TYPE "HMI Station: Wip Select: Screen"
   STRUCT
      animate : Array[0.."wipSelScrnObjCnt"] of Int;
      pbs : DWord;
      txt : Array[0.."wipSelScrnObjCnt"] of WString ["LONG_STRING_LENGTH"];
   END_STRUCT;
   // // txt[6] : wip select 00 label
   // // txt[7] : wip select 00 text
   // // txt[8] : wip select 01 label
   // // txt[9] : wip select 01 text
   // // txt[10] : wip select 02 label
   // // txt[11] : wip select 02 text
   // // txt[12] : wip select 03 label
   // // txt[13] : wip select 03 text
   // // txt[14] : wip select 04 label
   // // txt[15] : wip select 04 text
   // // txt[16] : wip select 05 label
   // // txt[17] : wip select 05 text
END_TYPE

TYPE "HMI Station: Template Screen"
   STRUCT
      animate : Array[0.."tmpltScrnObjCnt"] of Int;
      pb : DWord;
      text : Array[0.."tmpltScrnObjCnt"] of WString ["LONG_STRING_LENGTH"];
   END_STRUCT;
END_TYPE

// folder: KP8 Driver

TYPE "KP8 I/O Data"
   STRUCT
      input : Word;
      tempOut : DWord;
      finalOut : DWord;
   END_STRUCT;
END_TYPE

TYPE "KP8 Driver: Parameters: 1 Button"
   STRUCT
      activate : Bool;   // true = button on, flase = button off
      cOn1 : String[10];   // color when button is in pressed state. valid entries: 'red', 'green', 'blue', 'yellow', 'white', 'off'
      cOn2 : String[10];   // second flash color when button is pressed and flashing is enabled. valid entries: 'red', 'green', 'blue', 'yellow', 'white', 'off'
      cOff : String[10];   // color when button is in un-pressed state. valid entries: 'red', 'green', 'blue', 'yellow', 'white', 'off'
      flash : Bool;   // false = color 1, true = color 2. set to clock bit to flash at that rate
      group : Int;   // 0 disables. buttons in groups have a mutually exclusive 'on' state.
      mode : Bool;   // true = maintained, fales = momentary
   END_STRUCT;
END_TYPE

TYPE "KP8 Driver: Button States"
   STRUCT
      btn : Array[0..7] of Bool;
   END_STRUCT;
END_TYPE

TYPE "KP8 Driver: Parameters: 8 Buttons"
   STRUCT
      btn : Array[0..7] of "KP8 Driver: Parameters: 1 Button";
   END_STRUCT;
END_TYPE

TYPE "KP8 Driver: Feedback Data"
   STRUCT
      acutal : "KP8 Driver: Button States";
      falling : "KP8 Driver: Button States";
      rising : "KP8 Driver: Button States";
   END_STRUCT;
END_TYPE

// folder: Linked List

TYPE "Linked List: Node: Data"
   STRUCT
      place_holder : Int;
   END_STRUCT;
END_TYPE

TYPE "Linked List: Node: Meta"
   STRUCT
      key : DInt := -1;
      is_head : Bool;
      is_tail : Bool;
      next : DInt := -1;
   END_STRUCT;
END_TYPE

TYPE "Linked List: Node"
   STRUCT
      data : "Linked List: Node: Data";
      meta : "Linked List: Node: Meta";
   END_STRUCT;
END_TYPE

TYPE "Linked List: List"
   STRUCT
      me : Array[0.."LINKED_LIST_LENGTH"] of "Linked List: Node";
   END_STRUCT;
END_TYPE

TYPE "Linked List: Method Interface: Reset: In"
   STRUCT
      request : Bool;
   END_STRUCT;
END_TYPE

TYPE "Linked List: Method Interface: Reverse: Out"
   STRUCT
      done : Bool;
      error : Bool;
      error_message : String;
   END_STRUCT;
END_TYPE

TYPE "Linked List: Method Interface: Reverse: In"
   STRUCT
      request : Bool;
   END_STRUCT;
END_TYPE

TYPE "Linked List: Method Interface: Display: Out"
   STRUCT
      done : Bool;
      list : "Linked List: List";
   END_STRUCT;
END_TYPE

TYPE "Linked List: Method Interface: Display: In"
   STRUCT
      request : Bool;
   END_STRUCT;
END_TYPE

TYPE "Linked List: Method Interface: Search: Out"
   STRUCT
      done : Bool;
      error : Bool;
      error_message : String;
      found : Bool;
      not_found : Bool;
      returned_node : "Linked List: Node";
   END_STRUCT;
END_TYPE

TYPE "Linked List: Method Interface: Search: In"
   STRUCT
      data : "Linked List: Node: Data";
      request : Bool;
   END_STRUCT;
END_TYPE

TYPE "Linked List: Method Interface: Reset: Out"
   STRUCT
      done : Bool;
   END_STRUCT;
END_TYPE

TYPE "Linked List: Method Interface: Delete: Out"
   STRUCT
      done : Bool;
      error : Bool;
      error_message : String;
   END_STRUCT;
END_TYPE

TYPE "Linked List: Method Interface: Delete: In"
   STRUCT
      node : "Linked List: Node";   // key of node to be deleted
      request : Bool;
   END_STRUCT;
END_TYPE

TYPE "Linked List: Method Interface: Insert: Out"
   STRUCT
      done : Bool;
      error : Bool;
      error_message : String;
   END_STRUCT;
END_TYPE

TYPE "Linked List: Method Interface: Insert: In"
   STRUCT
      target_node : "Linked List: Node";   // key of node after which new node is to be inserted
      data : "Linked List: Node: Data";
      request : Bool;
   END_STRUCT;
END_TYPE

TYPE "Linked List: Method Interface: Append: In"
   STRUCT
      data : "Linked List: Node: Data";
      request : Bool;
   END_STRUCT;
END_TYPE

TYPE "Linked List: Method Interface: Append: Out"
   STRUCT
      done : Bool;
      error : Bool;
      error_message : String;
   END_STRUCT;
END_TYPE

TYPE "Linked List: Method Interface: Delete"
   STRUCT
      in : "Linked List: Method Interface: Delete: In";
      out : "Linked List: Method Interface: Delete: Out";
   END_STRUCT;
END_TYPE

TYPE "Linked List: Method Interface: Search"
   STRUCT
      in : "Linked List: Method Interface: Search: In";
      out : "Linked List: Method Interface: Search: Out";
   END_STRUCT;
END_TYPE

TYPE "Linked List: Method Interface: Insert"
   STRUCT
      in : "Linked List: Method Interface: Insert: In";
      out : "Linked List: Method Interface: Insert: Out";
   END_STRUCT;
END_TYPE

TYPE "Linked List: Method Interface: Append"
   STRUCT
      in : "Linked List: Method Interface: Append: In";
      out : "Linked List: Method Interface: Append: Out";
   END_STRUCT;
END_TYPE

TYPE "Linked List: Method Interface: Reverse"
   STRUCT
      in : "Linked List: Method Interface: Reverse: In";
      out : "Linked List: Method Interface: Reverse: Out";
   END_STRUCT;
END_TYPE

TYPE "Linked List: Method Interface: Display"
   STRUCT
      in : "Linked List: Method Interface: Display: In";
      out : "Linked List: Method Interface: Display: Out";
   END_STRUCT;
END_TYPE

TYPE "Linked List: Method Interface: Reset"
   STRUCT
      in : "Linked List: Method Interface: Reset: In";
      out : "Linked List: Method Interface: Reset: Out";
   END_STRUCT;
END_TYPE

TYPE "Linked List: Method Interface"
   STRUCT
      append : "Linked List: Method Interface: Append";   // adds node containing data specified to end of list
      delete : "Linked List: Method Interface: Delete";   // removes the specified node
      display : "Linked List: Method Interface: Display";
      insert : "Linked List: Method Interface: Insert";   // inserts node containing data specified after node specified
      reset : "Linked List: Method Interface: Reset";
      reverse : "Linked List: Method Interface: Reverse";
      search : "Linked List: Method Interface: Search";   // returns the specified node
   END_STRUCT;
END_TYPE

// folder: Settings Screen New Data

TYPE "Settings Screen: Processed Inputs"
   STRUCT
      assign : "Push Button Data: State Change Data";
      line_name : "State Changes: WString";
      dropzone : "State Changes: WString";
      total : "State Changes: Real";
      critical : "State Changes: Real";
      part_number_single : "State Changes: WString";
      part_number_double : "State Changes: WString";
   END_STRUCT;
END_TYPE

// folder: State Changes

TYPE "State Changes: Bool"
   STRUCT
      rising : Bool;   // also used when tracking value changes
      falling : Bool;
      actual : Bool;
   END_STRUCT;
END_TYPE

TYPE "State Changes: WString"
   STRUCT
      rising : Bool;
      falling : Bool;
      actual : WString;
   END_STRUCT;
END_TYPE

TYPE "State Changes: Int"
   STRUCT
      rising : Bool;
      falling : Bool;
      actual : Int;
   END_STRUCT;
END_TYPE

TYPE "State Changes: UInt"
   STRUCT
      rising : Bool;
      falling : Bool;
      actual : UInt;
   END_STRUCT;
END_TYPE

TYPE "State Changes: USInt"
   STRUCT
      rising : Bool;
      falling : Bool;
      actual : USInt;
   END_STRUCT;
END_TYPE

TYPE "State Changes: Real"
   STRUCT
      rising : Bool;
      falling : Bool;
      actual : Real;
   END_STRUCT;
END_TYPE

// folder: Station

TYPE "Station: All Stations"
   STRUCT
      stn : Array[0.."STATION_COUNT"] of "Station: Single Station";
   END_STRUCT;
END_TYPE

TYPE "Station: Wip: Wip Module"
   STRUCT
      ioData : "Station I/O Data";
      flags : "Station: Wip Flags";
      kp8Logical : "KP8 Driver: Feedback Data";
      orderState : Array[0.."STATION_BUTTON_COUNT"] of Int;
      pnCode : Array[0.."STATION_BUTTON_COUNT"] of DInt;
      timers : "Station: Timers";
      wip : "Station: Wip: Meta Data: Single";
   END_STRUCT;
END_TYPE

TYPE "Station: Order States"
   STRUCT
      btn : Array[0.."STATION_BUTTON_COUNT"] of Int;
   END_STRUCT;
END_TYPE

TYPE "Station: KP8 Config"
VERSION : 0.1
   STRUCT
      activate : Bool;
      colorOn1 : String[10];
      colorOn2 : String[10];
      colorOff : String[10];
      flash : Bool;
      group : Int;
      mode : Bool;
   END_STRUCT;
END_TYPE

TYPE "Station: PN Code"
   STRUCT
      btn : Array[0.."STATION_BUTTON_COUNT"] of DInt;
   END_STRUCT;
END_TYPE

TYPE "Station: Single Station"
   STRUCT
      flags : "Station: Flags";
      id : "Station: Id";
      kp8Config : "KP8 Driver: Parameters: 8 Buttons";
      kp8Physical : "KP8 Driver: Feedback Data";
      wipData : "Station: Wip: Meta Data: All";
      wipCmpts : "Station: Wip: Wip Module";
   END_STRUCT;
END_TYPE

TYPE "Station: Animations"
   STRUCT
      btn : Array[0.."STATION_BUTTON_COUNT"] of UInt;
   END_STRUCT;
END_TYPE

TYPE "Station Selection Change"
   STRUCT
      falling : Bool;
      rising : Bool;
      selection_change : Bool;
      station_index : Int := -1;
   END_STRUCT;
END_TYPE

TYPE "Station: Sim Data"
   STRUCT
      stn : Struct
         animate : USInt;
         label : WString[20];
      END_STRUCT;
      btn : Struct
         actuate : Byte;
         animate : Array[0..7] of USInt;
         labels : Array[0..7] of WString [4];
      END_STRUCT;
   END_STRUCT;
END_TYPE

TYPE "Station: Wip Flags"
   STRUCT
      clearWipRequest : Bool;   // set: after wip has been deselected for deselect interval; consumed:
      inSettingsScreen : Bool;   // set: Flags: HMI Warehouse; consumed: Settings; reset: Flags: HMI Warehouse
      whHmiOrdered : Bool;   // set: Flags: HMI Warehouse, set by user input; consumed: Order State: Enter Ordered; reset: Order State: Enter Ordered
      newPN : Bool;   // set: Flags: New PN Code; reset:
      pnGood : Array[0.."STATION_BUTTON_COUNT"] of Bool;
      resetStation : Bool;
      resetTimer : Array[0.."STATION_BUTTON_COUNT"] of Bool;
   END_STRUCT;
END_TYPE

TYPE "Station: ET200SP Comm Debug Data"
   STRUCT
      dismissPB : Bool;
      IM : "ET200SP: IM Data";
      DQ01 : "ET200SP: DQ Data";
      DQ02 : "ET200SP: DQ Data";
      DQ03 : "ET200SP: DQ Data";
      profinetName : Struct
         animate : USInt;
         label : WString[20];
      END_STRUCT;
      serverModule : "ET200SP: Server Module Data";
   END_STRUCT;
END_TYPE

TYPE "Station: KP8 Comm Debug Data"
   STRUCT
      dismissPB : Bool;
      profinetName : Struct
         animate : USInt;
         label : WString[20];
      END_STRUCT;
      stencilBackground : USInt;
      X1P1 : Struct
         transmit : USInt;
         receive : USInt;
      END_STRUCT;
      X1P2 : Struct
         transmit : USInt;
         receive : USInt;
      END_STRUCT;
   END_STRUCT;
END_TYPE

TYPE "Station: Timers"
   STRUCT
      elapsed : Array[0.."STATION_BUTTON_COUNT"] of Real;   // time (s) that a part number has been requested
      ptAllotted : Array[0.."STATION_BUTTON_COUNT"] of Real;   // time (s) before a part request is considered over-due
      ptCritical : Array[0.."STATION_BUTTON_COUNT"] of Real;   // time (s) before a part request is considered critical
      remaining : Array[0.."STATION_BUTTON_COUNT"] of Real;   // request allotted - elapsed
      wsAllotted : Real := 10.0;   // time (s) before a selected wip is counted as being selected
      wsElapsed : Real;   // time (s) a wip has been selected
      wsRemaining : Real;   // wip select allotted - selected
      wdsAllotted : Real := 10.0;   // time (s) before a deselected wip's requests are cleared from the part request table
      wdsElapsed : Real;   // time (s) a wip has been deselected
      wdsRemaining : Real;   // wip deselect allotted - selected
   END_STRUCT;
END_TYPE

TYPE "Station: Wip: Meta Data: Single"
   STRUCT
      code : DInt := -1;   // builds station name from libraries
      useCount : DInt;   // number of times station selected for longer than lower dwell limit
   END_STRUCT;
END_TYPE

TYPE "Station: Flags"
   STRUCT
      stateTransition : Array[0.."STATION_BUTTON_COUNT"] of Bool;
      wipSwapped : Bool;
   END_STRUCT;
END_TYPE

TYPE "Station: Id"
   STRUCT
      dropZone : USInt;
      lineName : WString["SHORT_STRING_LENGTH"];
   END_STRUCT;
END_TYPE

TYPE "Station I/O Data"
   STRUCT
      kp8 : "KP8 I/O Data";
      stkLight : DWord;
   END_STRUCT;
END_TYPE

TYPE "Station: Wip: Meta Data: All"
   STRUCT
      code : DInt := -1;   // wip label library code for currently selected wip
      count : DInt;   // number of wips in this station
      index : DInt := -1;   // index in saved wip array of currently selected wip
   END_STRUCT;
END_TYPE

// folder: (top level)

DATA_BLOCK "EMP IDB"   // DB1
{ S7_Optimized_Access := 'TRUE' }
VERSION : 0.1
// stored: InstanceOfName EMP
"EMP"
BEGIN
   "inst HMI Station"."inst HMI Station: Wip Selection".rowIndicies[1] := 1;
   "inst HMI Station"."inst HMI Station: Wip Selection".rowIndicies[2] := 2;
   "inst HMI Station"."inst HMI Station: Wip Selection".rowIndicies[3] := 3;
   "inst HMI Station"."inst HMI Station: Wip Selection".rowIndicies[4] := 4;
   "inst HMI Station"."inst HMI Station: Wip Selection".rowIndicies[5] := 5;
END_DATA_BLOCK

DATA_BLOCK "Debug"   // DB7
{ S7_Optimized_Access := 'TRUE' }
VERSION : 0.1
   VAR
      search_term : WString;
      index : Int;
      test : Bool;
      rep : Int;
      "rep*len" : Int;
      "i+rep*len" : Int;
   END_VAR
BEGIN
END_DATA_BLOCK

// folder: From Excel

DATA_BLOCK "From Excel: Codes"   // DB12
{ S7_Optimized_Access := 'TRUE' }
VERSION : 0.1
BEGIN
   kp8Stns[0].pnCode[0] := 0;
   kp8Stns[0].pnCode[1] := 0;
   kp8Stns[0].pnCode[2] := 0;
   kp8Stns[0].pnCode[3] := 172000;
   kp8Stns[0].pnCode[4] := 0;
   kp8Stns[0].pnCode[5] := 0;
   kp8Stns[0].pnCode[6] := 0;
   kp8Stns[0].pnCode[7] := 168000;
   kp8Stns[1].pnCode[0] := 0;
   kp8Stns[1].pnCode[1] := 0;
   kp8Stns[1].pnCode[2] := 183000;
   kp8Stns[1].pnCode[3] := 209000;
   kp8Stns[1].pnCode[4] := 0;
   kp8Stns[1].pnCode[5] := 0;
   kp8Stns[1].pnCode[6] := 180000;
   kp8Stns[1].pnCode[7] := 166000;
   kp8Stns[2].pnCode[0] := 0;
   kp8Stns[2].pnCode[1] := 182000;
   kp8Stns[2].pnCode[2] := 181000;
   kp8Stns[2].pnCode[3] := 215000;
   kp8Stns[2].pnCode[4] := 0;
   kp8Stns[2].pnCode[5] := 184000;
   kp8Stns[2].pnCode[6] := 216000;
   kp8Stns[2].pnCode[7] := 214000;
   kp8Stns[3].pnCode[0] := 0;
   kp8Stns[3].pnCode[1] := 192000;
   kp8Stns[3].pnCode[2] := 191000;
   kp8Stns[3].pnCode[3] := 188000;
   kp8Stns[3].pnCode[4] := 0;
   kp8Stns[3].pnCode[5] := 190000;
   kp8Stns[3].pnCode[6] := 187000;
   kp8Stns[3].pnCode[7] := 189000;
   kp8Stns[4].pnCode[0] := 0;
   kp8Stns[4].pnCode[1] := 0;
   kp8Stns[4].pnCode[2] := 0;
   kp8Stns[4].pnCode[3] := 0;
   kp8Stns[4].pnCode[4] := 0;
   kp8Stns[4].pnCode[5] := 0;
   kp8Stns[4].pnCode[6] := 0;
   kp8Stns[4].pnCode[7] := 194000;
   kp8Stns[5].pnCode[0] := 0;
   kp8Stns[5].pnCode[1] := 193000;
   kp8Stns[5].pnCode[2] := 195000;
   kp8Stns[5].pnCode[3] := 176000;
   kp8Stns[5].pnCode[4] := 0;
   kp8Stns[5].pnCode[5] := 196000;
   kp8Stns[5].pnCode[6] := 177000;
   kp8Stns[5].pnCode[7] := 175000;
   kp8Stns[6].pnCode[0] := 0;
   kp8Stns[6].pnCode[1] := 208000;
   kp8Stns[6].pnCode[2] := 207000;
   kp8Stns[6].pnCode[3] := 210000;
   kp8Stns[6].pnCode[4] := 0;
   kp8Stns[6].pnCode[5] := 211000;
   kp8Stns[6].pnCode[6] := 206000;
   kp8Stns[6].pnCode[7] := 205000;
   kp8Stns[7].pnCode[0] := 0;
   kp8Stns[7].pnCode[1] := 0;
   kp8Stns[7].pnCode[2] := 0;
   kp8Stns[7].pnCode[3] := 174000;
   kp8Stns[7].pnCode[4] := 0;
   kp8Stns[7].pnCode[5] := 0;
   kp8Stns[7].pnCode[6] := 167000;
   kp8Stns[7].pnCode[7] := 169000;
   kp8Stns[8].pnCode[0] := 0;
   kp8Stns[8].pnCode[1] := 0;
   kp8Stns[8].pnCode[2] := 0;
   kp8Stns[8].pnCode[3] := 204000;
   kp8Stns[8].pnCode[4] := 0;
   kp8Stns[8].pnCode[5] := 0;
   kp8Stns[8].pnCode[6] := 173000;
   kp8Stns[8].pnCode[7] := 186000;
   kp8Stns[9].pnCode[0] := 0;
   kp8Stns[9].pnCode[1] := 0;
   kp8Stns[9].pnCode[2] := 0;
   kp8Stns[9].pnCode[3] := 213000;
   kp8Stns[9].pnCode[4] := 0;
   kp8Stns[9].pnCode[5] := 0;
   kp8Stns[9].pnCode[6] := 0;
   kp8Stns[9].pnCode[7] := 212000;
   kp8Stns[10].pnCode[0] := 0;
   kp8Stns[10].pnCode[1] := 0;
   kp8Stns[10].pnCode[2] := 0;
   kp8Stns[10].pnCode[3] := 170000;
   kp8Stns[10].pnCode[4] := 0;
   kp8Stns[10].pnCode[5] := 0;
   kp8Stns[10].pnCode[6] := 242000;
   kp8Stns[10].pnCode[7] := 171000;
   kp8Stns[11].pnCode[0] := 0;
   kp8Stns[11].pnCode[1] := 0;
   kp8Stns[11].pnCode[2] := 0;
   kp8Stns[11].pnCode[3] := 77000;
   kp8Stns[11].pnCode[4] := 0;
   kp8Stns[11].pnCode[5] := 0;
   kp8Stns[11].pnCode[6] := 65000;
   kp8Stns[11].pnCode[7] := 20000;
   kp8Stns[12].pnCode[0] := 0;
   kp8Stns[12].pnCode[1] := 80000;
   kp8Stns[12].pnCode[2] := 86000;
   kp8Stns[12].pnCode[3] := 59000;
   kp8Stns[12].pnCode[4] := 0;
   kp8Stns[12].pnCode[5] := 79000;
   kp8Stns[12].pnCode[6] := 55000;
   kp8Stns[12].pnCode[7] := 54000;
   kp8Stns[13].pnCode[0] := 0;
   kp8Stns[13].pnCode[1] := 0;
   kp8Stns[13].pnCode[2] := 69000;
   kp8Stns[13].pnCode[3] := 89000;
   kp8Stns[13].pnCode[4] := 0;
   kp8Stns[13].pnCode[5] := 0;
   kp8Stns[13].pnCode[6] := 90000;
   kp8Stns[13].pnCode[7] := 88000;
   kp8Stns[14].pnCode[0] := 0;
   kp8Stns[14].pnCode[1] := 0;
   kp8Stns[14].pnCode[2] := 64000;
   kp8Stns[14].pnCode[3] := 87000;
   kp8Stns[14].pnCode[4] := 0;
   kp8Stns[14].pnCode[5] := 63000;
   kp8Stns[14].pnCode[6] := 82000;
   kp8Stns[14].pnCode[7] := 62000;
   kp8Stns[15].pnCode[0] := 0;
   kp8Stns[15].pnCode[1] := 49000;
   kp8Stns[15].pnCode[2] := 76000;
   kp8Stns[15].pnCode[3] := 28000;
   kp8Stns[15].pnCode[4] := 0;
   kp8Stns[15].pnCode[5] := 81000;
   kp8Stns[15].pnCode[6] := 68000;
   kp8Stns[15].pnCode[7] := 74000;
   kp8Stns[16].pnCode[0] := 0;
   kp8Stns[16].pnCode[1] := 0;
   kp8Stns[16].pnCode[2] := 0;
   kp8Stns[16].pnCode[3] := 91000;
   kp8Stns[16].pnCode[4] := 0;
   kp8Stns[16].pnCode[5] := 0;
   kp8Stns[16].pnCode[6] := 93000;
   kp8Stns[16].pnCode[7] := 94067;
   kp8Stns[17].pnCode[0] := 0;
   kp8Stns[17].pnCode[1] := 0;
   kp8Stns[17].pnCode[2] := 83000;
   kp8Stns[17].pnCode[3] := 34000;
   kp8Stns[17].pnCode[4] := 0;
   kp8Stns[17].pnCode[5] := 0;
   kp8Stns[17].pnCode[6] := 75000;
   kp8Stns[17].pnCode[7] := 29000;
   kp8Stns[18].pnCode[0] := 0;
   kp8Stns[18].pnCode[1] := 0;
   kp8Stns[18].pnCode[2] := 0;
   kp8Stns[18].pnCode[3] := 92066;
   kp8Stns[18].pnCode[4] := 0;
   kp8Stns[18].pnCode[5] := 0;
   kp8Stns[18].pnCode[6] := 96026;
   kp8Stns[18].pnCode[7] := 95000;
   kp8Stns[19].pnCode[0] := 0;
   kp8Stns[19].pnCode[1] := 78000;
   kp8Stns[19].pnCode[2] := 85000;
   kp8Stns[19].pnCode[3] := 21000;
   kp8Stns[19].pnCode[4] := 0;
   kp8Stns[19].pnCode[5] := 97000;
   kp8Stns[19].pnCode[6] := 60000;
   kp8Stns[19].pnCode[7] := 48000;
   kp8Stns[20].pnCode[0] := 0;
   kp8Stns[20].pnCode[1] := 0;
   kp8Stns[20].pnCode[2] := 0;
   kp8Stns[20].pnCode[3] := 0;
   kp8Stns[20].pnCode[4] := 0;
   kp8Stns[20].pnCode[5] := 0;
   kp8Stns[20].pnCode[6] := 0;
   kp8Stns[20].pnCode[7] := 244000;
   kp8Stns[21].pnCode[0] := 0;
   kp8Stns[21].pnCode[1] := 0;
   kp8Stns[21].pnCode[2] := 0;
   kp8Stns[21].pnCode[3] := 245000;
   kp8Stns[21].pnCode[4] := 0;
   kp8Stns[21].pnCode[5] := 0;
   kp8Stns[21].pnCode[6] := 0;
   kp8Stns[21].pnCode[7] := 11000;
   kp8Stns[22].pnCode[0] := 0;
   kp8Stns[22].pnCode[1] := 0;
   kp8Stns[22].pnCode[2] := 0;
   kp8Stns[22].pnCode[3] := 22000;
   kp8Stns[22].pnCode[4] := 0;
   kp8Stns[22].pnCode[5] := 0;
   kp8Stns[22].pnCode[6] := 46000;
   kp8Stns[22].pnCode[7] := 61000;
   kp8Stns[23].pnCode[0] := 0;
   kp8Stns[23].pnCode[1] := 0;
   kp8Stns[23].pnCode[2] := 0;
   kp8Stns[23].pnCode[3] := 0;
   kp8Stns[23].pnCode[4] := 0;
   kp8Stns[23].pnCode[5] := 0;
   kp8Stns[23].pnCode[6] := 0;
   kp8Stns[23].pnCode[7] := 12000;
   kp8Stns[24].pnCode[0] := 0;
   kp8Stns[24].pnCode[1] := 0;
   kp8Stns[24].pnCode[2] := 0;
   kp8Stns[24].pnCode[3] := 0;
   kp8Stns[24].pnCode[4] := 0;
   kp8Stns[24].pnCode[5] := 0;
   kp8Stns[24].pnCode[6] := 0;
   kp8Stns[24].pnCode[7] := 27000;
   kp8Stns[25].pnCode[0] := 0;
   kp8Stns[25].pnCode[1] := 0;
   kp8Stns[25].pnCode[2] := 0;
   kp8Stns[25].pnCode[3] := 0;
   kp8Stns[25].pnCode[4] := 0;
   kp8Stns[25].pnCode[5] := 0;
   kp8Stns[25].pnCode[6] := 0;
   kp8Stns[25].pnCode[7] := 56000;
   hmiStns[0].wip[0].wipCode := 6027;
   hmiStns[0].wip[0].pnCode[0] := 0;
   hmiStns[0].wip[0].pnCode[1] := 243000;
   hmiStns[0].wip[0].pnCode[2] := 19000;
   hmiStns[0].wip[0].pnCode[3] := 0;
   hmiStns[0].wip[0].pnCode[4] := 0;
   hmiStns[0].wip[0].pnCode[5] := 0;
   hmiStns[0].wip[0].pnCode[6] := 25000;
   hmiStns[0].wip[0].pnCode[7] := 18000;
   hmiStns[0].wip[1].wipCode := 9007;
   hmiStns[0].wip[1].pnCode[0] := 0;
   hmiStns[0].wip[1].pnCode[1] := 243000;
   hmiStns[0].wip[1].pnCode[2] := 37000;
   hmiStns[0].wip[1].pnCode[3] := 0;
   hmiStns[0].wip[1].pnCode[4] := 0;
   hmiStns[0].wip[1].pnCode[5] := 0;
   hmiStns[0].wip[1].pnCode[6] := 35000;
   hmiStns[0].wip[1].pnCode[7] := 36000;
   hmiStns[0].wip[2].wipCode := 10030;
   hmiStns[0].wip[2].pnCode[0] := 0;
   hmiStns[0].wip[2].pnCode[1] := 243000;
   hmiStns[0].wip[2].pnCode[2] := 40000;
   hmiStns[0].wip[2].pnCode[3] := 0;
   hmiStns[0].wip[2].pnCode[4] := 0;
   hmiStns[0].wip[2].pnCode[5] := 0;
   hmiStns[0].wip[2].pnCode[6] := 38000;
   hmiStns[0].wip[2].pnCode[7] := 39000;
   hmiStns[0].wip[3].wipCode := 11056;
   hmiStns[0].wip[3].pnCode[0] := 0;
   hmiStns[0].wip[3].pnCode[1] := 243000;
   hmiStns[0].wip[3].pnCode[2] := 47000;
   hmiStns[0].wip[3].pnCode[3] := 13000;
   hmiStns[0].wip[3].pnCode[4] := 0;
   hmiStns[0].wip[3].pnCode[5] := 14000;
   hmiStns[0].wip[3].pnCode[6] := 41000;
   hmiStns[0].wip[3].pnCode[7] := 32000;
   hmiStns[0].wip[4].wipCode := 12008;
   hmiStns[0].wip[4].pnCode[0] := 0;
   hmiStns[0].wip[4].pnCode[1] := 243000;
   hmiStns[0].wip[4].pnCode[2] := 45000;
   hmiStns[0].wip[4].pnCode[3] := 0;
   hmiStns[0].wip[4].pnCode[4] := 0;
   hmiStns[0].wip[4].pnCode[5] := 0;
   hmiStns[0].wip[4].pnCode[6] := 35000;
   hmiStns[0].wip[4].pnCode[7] := 36000;
   hmiStns[0].wip[5].wipCode := 13060;
   hmiStns[0].wip[5].pnCode[0] := 0;
   hmiStns[0].wip[5].pnCode[1] := 243000;
   hmiStns[0].wip[5].pnCode[2] := 37000;
   hmiStns[0].wip[5].pnCode[3] := 0;
   hmiStns[0].wip[5].pnCode[4] := 0;
   hmiStns[0].wip[5].pnCode[5] := 0;
   hmiStns[0].wip[5].pnCode[6] := 42000;
   hmiStns[0].wip[5].pnCode[7] := 36000;
   hmiStns[0].wip[6].wipCode := 14061;
   hmiStns[0].wip[6].pnCode[0] := 0;
   hmiStns[0].wip[6].pnCode[1] := 243000;
   hmiStns[0].wip[6].pnCode[2] := 45000;
   hmiStns[0].wip[6].pnCode[3] := 0;
   hmiStns[0].wip[6].pnCode[4] := 0;
   hmiStns[0].wip[6].pnCode[5] := 0;
   hmiStns[0].wip[6].pnCode[6] := 42000;
   hmiStns[0].wip[6].pnCode[7] := 36000;
   hmiStns[0].wip[7].wipCode := 15030;
   hmiStns[0].wip[7].pnCode[0] := 0;
   hmiStns[0].wip[7].pnCode[1] := 243000;
   hmiStns[0].wip[7].pnCode[2] := 43000;
   hmiStns[0].wip[7].pnCode[3] := 0;
   hmiStns[0].wip[7].pnCode[4] := 0;
   hmiStns[0].wip[7].pnCode[5] := 0;
   hmiStns[0].wip[7].pnCode[6] := 38000;
   hmiStns[0].wip[7].pnCode[7] := 44000;
   hmiStns[0].wip[8].wipCode := 16024;
   hmiStns[0].wip[8].pnCode[0] := 0;
   hmiStns[0].wip[8].pnCode[1] := 243000;
   hmiStns[0].wip[8].pnCode[2] := 51000;
   hmiStns[0].wip[8].pnCode[3] := 0;
   hmiStns[0].wip[8].pnCode[4] := 0;
   hmiStns[0].wip[8].pnCode[5] := 0;
   hmiStns[0].wip[8].pnCode[6] := 25000;
   hmiStns[0].wip[8].pnCode[7] := 18000;
   hmiStns[0].wip[9].wipCode := 17009;
   hmiStns[0].wip[9].pnCode[0] := 0;
   hmiStns[0].wip[9].pnCode[1] := 243000;
   hmiStns[0].wip[9].pnCode[2] := 52000;
   hmiStns[0].wip[9].pnCode[3] := 0;
   hmiStns[0].wip[9].pnCode[4] := 0;
   hmiStns[0].wip[9].pnCode[5] := 0;
   hmiStns[0].wip[9].pnCode[6] := 31000;
   hmiStns[0].wip[9].pnCode[7] := 73000;
   hmiStns[0].wip[10].wipCode := 19031;
   hmiStns[0].wip[10].pnCode[0] := 0;
   hmiStns[0].wip[10].pnCode[1] := 243000;
   hmiStns[0].wip[10].pnCode[2] := 53000;
   hmiStns[0].wip[10].pnCode[3] := 0;
   hmiStns[0].wip[10].pnCode[4] := 0;
   hmiStns[0].wip[10].pnCode[5] := 0;
   hmiStns[0].wip[10].pnCode[6] := 31000;
   hmiStns[0].wip[10].pnCode[7] := 71000;
   hmiStns[0].wip[11].wipCode := 21028;
   hmiStns[0].wip[11].pnCode[0] := 0;
   hmiStns[0].wip[11].pnCode[1] := 243000;
   hmiStns[0].wip[11].pnCode[2] := 57000;
   hmiStns[0].wip[11].pnCode[3] := 0;
   hmiStns[0].wip[11].pnCode[4] := 0;
   hmiStns[0].wip[11].pnCode[5] := 0;
   hmiStns[0].wip[11].pnCode[6] := 25000;
   hmiStns[0].wip[11].pnCode[7] := 18000;
   hmiStns[0].wip[12].wipCode := 22008;
   hmiStns[0].wip[12].pnCode[0] := 0;
   hmiStns[0].wip[12].pnCode[1] := 243000;
   hmiStns[0].wip[12].pnCode[2] := 84000;
   hmiStns[0].wip[12].pnCode[3] := 0;
   hmiStns[0].wip[12].pnCode[4] := 0;
   hmiStns[0].wip[12].pnCode[5] := 0;
   hmiStns[0].wip[12].pnCode[6] := 31000;
   hmiStns[0].wip[12].pnCode[7] := 71000;
   hmiStns[0].wip[13].wipCode := 24029;
   hmiStns[0].wip[13].pnCode[0] := 0;
   hmiStns[0].wip[13].pnCode[1] := 243000;
   hmiStns[0].wip[13].pnCode[2] := 98000;
   hmiStns[0].wip[13].pnCode[3] := 0;
   hmiStns[0].wip[13].pnCode[4] := 0;
   hmiStns[0].wip[13].pnCode[5] := 0;
   hmiStns[0].wip[13].pnCode[6] := 38000;
   hmiStns[0].wip[13].pnCode[7] := 44000;
   hmiStns[0].wip[14].wipCode := 25025;
   hmiStns[0].wip[14].pnCode[0] := 0;
   hmiStns[0].wip[14].pnCode[1] := 243000;
   hmiStns[0].wip[14].pnCode[2] := 99000;
   hmiStns[0].wip[14].pnCode[3] := 0;
   hmiStns[0].wip[14].pnCode[4] := 0;
   hmiStns[0].wip[14].pnCode[5] := 0;
   hmiStns[0].wip[14].pnCode[6] := 42000;
   hmiStns[0].wip[14].pnCode[7] := 36000;
   hmiStns[0].wip[15].wipCode := 26026;
   hmiStns[0].wip[15].pnCode[0] := 0;
   hmiStns[0].wip[15].pnCode[1] := 243000;
   hmiStns[0].wip[15].pnCode[2] := 99000;
   hmiStns[0].wip[15].pnCode[3] := 0;
   hmiStns[0].wip[15].pnCode[4] := 0;
   hmiStns[0].wip[15].pnCode[5] := 0;
   hmiStns[0].wip[15].pnCode[6] := 35000;
   hmiStns[0].wip[15].pnCode[7] := 36000;
   hmiStns[0].wip[16].wipCode := 69063;
   hmiStns[0].wip[16].pnCode[0] := 0;
   hmiStns[0].wip[16].pnCode[1] := 243000;
   hmiStns[0].wip[16].pnCode[2] := 217000;
   hmiStns[0].wip[16].pnCode[3] := 0;
   hmiStns[0].wip[16].pnCode[4] := 0;
   hmiStns[0].wip[16].pnCode[5] := 0;
   hmiStns[0].wip[16].pnCode[6] := 218000;
   hmiStns[0].wip[16].pnCode[7] := 223000;
   hmiStns[0].wip[17].wipCode := 71000;
   hmiStns[0].wip[17].pnCode[0] := 0;
   hmiStns[0].wip[17].pnCode[1] := 243000;
   hmiStns[0].wip[17].pnCode[2] := 197000;
   hmiStns[0].wip[17].pnCode[3] := 0;
   hmiStns[0].wip[17].pnCode[4] := 0;
   hmiStns[0].wip[17].pnCode[5] := 0;
   hmiStns[0].wip[17].pnCode[6] := 219000;
   hmiStns[0].wip[17].pnCode[7] := 222000;
   hmiStns[0].wip[18].wipCode := 72023;
   hmiStns[0].wip[18].pnCode[0] := 0;
   hmiStns[0].wip[18].pnCode[1] := 243000;
   hmiStns[0].wip[18].pnCode[2] := 198000;
   hmiStns[0].wip[18].pnCode[3] := 0;
   hmiStns[0].wip[18].pnCode[4] := 0;
   hmiStns[0].wip[18].pnCode[5] := 0;
   hmiStns[0].wip[18].pnCode[6] := 218000;
   hmiStns[0].wip[18].pnCode[7] := 223000;
   hmiStns[0].wip[19].wipCode := 73064;
   hmiStns[0].wip[19].pnCode[0] := 0;
   hmiStns[0].wip[19].pnCode[1] := 243000;
   hmiStns[0].wip[19].pnCode[2] := 224000;
   hmiStns[0].wip[19].pnCode[3] := 0;
   hmiStns[0].wip[19].pnCode[4] := 0;
   hmiStns[0].wip[19].pnCode[5] := 0;
   hmiStns[0].wip[19].pnCode[6] := 225000;
   hmiStns[0].wip[19].pnCode[7] := 226000;
   hmiStns[0].wip[20].wipCode := 5009;
   hmiStns[0].wip[20].pnCode[0] := 0;
   hmiStns[0].wip[20].pnCode[1] := 243000;
   hmiStns[0].wip[20].pnCode[2] := 17000;
   hmiStns[0].wip[20].pnCode[3] := 0;
   hmiStns[0].wip[20].pnCode[4] := 0;
   hmiStns[0].wip[20].pnCode[5] := 0;
   hmiStns[0].wip[20].pnCode[6] := 24000;
   hmiStns[0].wip[20].pnCode[7] := 16000;
   hmiStns[0].wip[21].wipCode := 7031;
   hmiStns[0].wip[21].pnCode[0] := 0;
   hmiStns[0].wip[21].pnCode[1] := 243000;
   hmiStns[0].wip[21].pnCode[2] := 0;
   hmiStns[0].wip[21].pnCode[3] := 31000;
   hmiStns[0].wip[21].pnCode[4] := 0;
   hmiStns[0].wip[21].pnCode[5] := 0;
   hmiStns[0].wip[21].pnCode[6] := 50000;
   hmiStns[0].wip[21].pnCode[7] := 30000;
   hmiStns[0].wip[22].wipCode := 74011;
   hmiStns[0].wip[22].pnCode[0] := 0;
   hmiStns[0].wip[22].pnCode[1] := 243000;
   hmiStns[0].wip[22].pnCode[2] := 0;
   hmiStns[0].wip[22].pnCode[3] := 219000;
   hmiStns[0].wip[22].pnCode[4] := 0;
   hmiStns[0].wip[22].pnCode[5] := 0;
   hmiStns[0].wip[22].pnCode[6] := 221000;
   hmiStns[0].wip[22].pnCode[7] := 222000;
   hmiStns[0].wip[23].wipCode := 70010;
   hmiStns[0].wip[23].pnCode[0] := 0;
   hmiStns[0].wip[23].pnCode[1] := 243000;
   hmiStns[0].wip[23].pnCode[2] := 220000;
   hmiStns[0].wip[23].pnCode[3] := 0;
   hmiStns[0].wip[23].pnCode[4] := 0;
   hmiStns[0].wip[23].pnCode[5] := 0;
   hmiStns[0].wip[23].pnCode[6] := 219000;
   hmiStns[0].wip[23].pnCode[7] := 222000;
   hmiStns[0].wip[24].wipCode := -1;
   hmiStns[0].wip[24].pnCode[0] := 0;
   hmiStns[0].wip[24].pnCode[1] := 0;
   hmiStns[0].wip[24].pnCode[2] := 0;
   hmiStns[0].wip[24].pnCode[3] := 0;
   hmiStns[0].wip[24].pnCode[4] := 0;
   hmiStns[0].wip[24].pnCode[5] := 0;
   hmiStns[0].wip[24].pnCode[6] := 0;
   hmiStns[0].wip[24].pnCode[7] := 0;
   hmiStns[0].wip[25].wipCode := -1;
   hmiStns[0].wip[25].pnCode[0] := 0;
   hmiStns[0].wip[25].pnCode[1] := 0;
   hmiStns[0].wip[25].pnCode[2] := 0;
   hmiStns[0].wip[25].pnCode[3] := 0;
   hmiStns[0].wip[25].pnCode[4] := 0;
   hmiStns[0].wip[25].pnCode[5] := 0;
   hmiStns[0].wip[25].pnCode[6] := 0;
   hmiStns[0].wip[25].pnCode[7] := 0;
   hmiStns[0].wip[26].wipCode := -1;
   hmiStns[0].wip[26].pnCode[0] := 0;
   hmiStns[0].wip[26].pnCode[1] := 0;
   hmiStns[0].wip[26].pnCode[2] := 0;
   hmiStns[0].wip[26].pnCode[3] := 0;
   hmiStns[0].wip[26].pnCode[4] := 0;
   hmiStns[0].wip[26].pnCode[5] := 0;
   hmiStns[0].wip[26].pnCode[6] := 0;
   hmiStns[0].wip[26].pnCode[7] := 0;
   hmiStns[0].wip[27].wipCode := -1;
   hmiStns[0].wip[27].pnCode[0] := 0;
   hmiStns[0].wip[27].pnCode[1] := 0;
   hmiStns[0].wip[27].pnCode[2] := 0;
   hmiStns[0].wip[27].pnCode[3] := 0;
   hmiStns[0].wip[27].pnCode[4] := 0;
   hmiStns[0].wip[27].pnCode[5] := 0;
   hmiStns[0].wip[27].pnCode[6] := 0;
   hmiStns[0].wip[27].pnCode[7] := 0;
   hmiStns[0].wip[28].wipCode := -1;
   hmiStns[0].wip[28].pnCode[0] := 0;
   hmiStns[0].wip[28].pnCode[1] := 0;
   hmiStns[0].wip[28].pnCode[2] := 0;
   hmiStns[0].wip[28].pnCode[3] := 0;
   hmiStns[0].wip[28].pnCode[4] := 0;
   hmiStns[0].wip[28].pnCode[5] := 0;
   hmiStns[0].wip[28].pnCode[6] := 0;
   hmiStns[0].wip[28].pnCode[7] := 0;
   hmiStns[0].wip[29].wipCode := -1;
   hmiStns[0].wip[29].pnCode[0] := 0;
   hmiStns[0].wip[29].pnCode[1] := 0;
   hmiStns[0].wip[29].pnCode[2] := 0;
   hmiStns[0].wip[29].pnCode[3] := 0;
   hmiStns[0].wip[29].pnCode[4] := 0;
   hmiStns[0].wip[29].pnCode[5] := 0;
   hmiStns[0].wip[29].pnCode[6] := 0;
   hmiStns[0].wip[29].pnCode[7] := 0;
   hmiStns[0].wip[30].wipCode := -1;
   hmiStns[0].wip[30].pnCode[0] := 0;
   hmiStns[0].wip[30].pnCode[1] := 0;
   hmiStns[0].wip[30].pnCode[2] := 0;
   hmiStns[0].wip[30].pnCode[3] := 0;
   hmiStns[0].wip[30].pnCode[4] := 0;
   hmiStns[0].wip[30].pnCode[5] := 0;
   hmiStns[0].wip[30].pnCode[6] := 0;
   hmiStns[0].wip[30].pnCode[7] := 0;
   hmiStns[0].wip[31].wipCode := -1;
   hmiStns[0].wip[31].pnCode[0] := 0;
   hmiStns[0].wip[31].pnCode[1] := 0;
   hmiStns[0].wip[31].pnCode[2] := 0;
   hmiStns[0].wip[31].pnCode[3] := 0;
   hmiStns[0].wip[31].pnCode[4] := 0;
   hmiStns[0].wip[31].pnCode[5] := 0;
   hmiStns[0].wip[31].pnCode[6] := 0;
   hmiStns[0].wip[31].pnCode[7] := 0;
   hmiStns[0].wip[32].wipCode := -1;
   hmiStns[0].wip[32].pnCode[0] := 0;
   hmiStns[0].wip[32].pnCode[1] := 0;
   hmiStns[0].wip[32].pnCode[2] := 0;
   hmiStns[0].wip[32].pnCode[3] := 0;
   hmiStns[0].wip[32].pnCode[4] := 0;
   hmiStns[0].wip[32].pnCode[5] := 0;
   hmiStns[0].wip[32].pnCode[6] := 0;
   hmiStns[0].wip[32].pnCode[7] := 0;
   hmiStns[0].wip[33].wipCode := -1;
   hmiStns[0].wip[33].pnCode[0] := 0;
   hmiStns[0].wip[33].pnCode[1] := 0;
   hmiStns[0].wip[33].pnCode[2] := 0;
   hmiStns[0].wip[33].pnCode[3] := 0;
   hmiStns[0].wip[33].pnCode[4] := 0;
   hmiStns[0].wip[33].pnCode[5] := 0;
   hmiStns[0].wip[33].pnCode[6] := 0;
   hmiStns[0].wip[33].pnCode[7] := 0;
   hmiStns[0].wip[34].wipCode := -1;
   hmiStns[0].wip[34].pnCode[0] := 0;
   hmiStns[0].wip[34].pnCode[1] := 0;
   hmiStns[0].wip[34].pnCode[2] := 0;
   hmiStns[0].wip[34].pnCode[3] := 0;